(* CODESYS project CanOpen.project (continued)
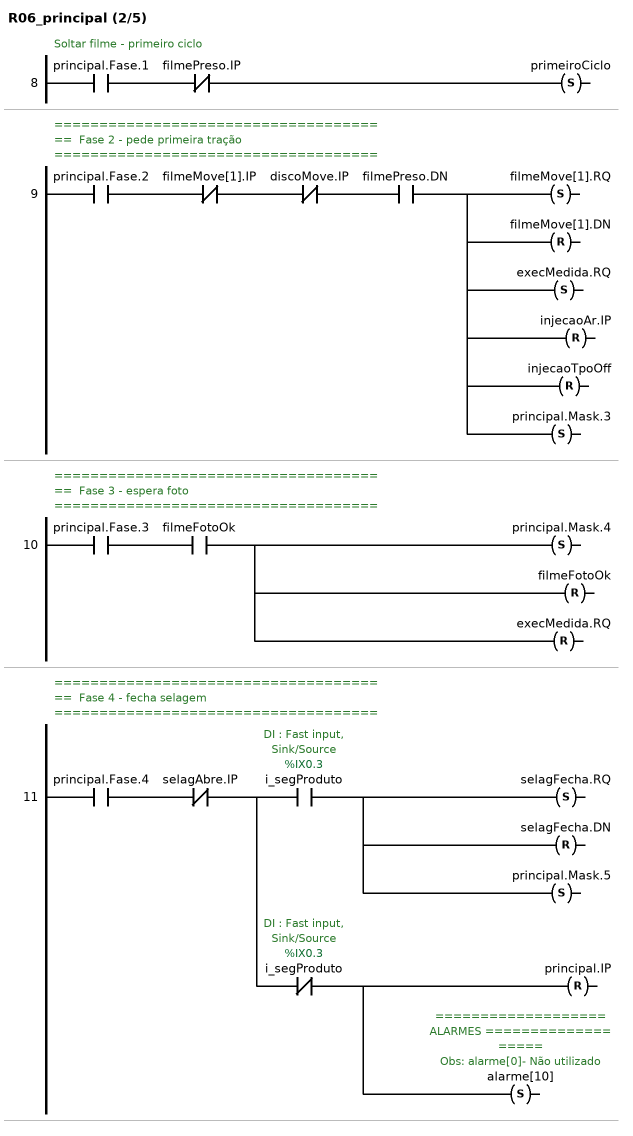
// NETWORK 8
// Soltar filme - primeiro ciclo
primeiroCiclo S= principal.Fase.1 AND NOT filmePreso.IP;

// NETWORK 9
// ====================================
// ==  Fase 2 - pede primeira tração
// ====================================
_w6 := principal.Fase.2 AND NOT filmeMove[1].IP AND NOT discoMove.IP AND filmePreso.DN;
filmeMove[1].RQ S= _w6;
filmeMove[1].DN R= _w6;
execMedida.RQ S= _w6;
injecaoAr.IP R= _w6;
injecaoTpoOff R= _w6;
principal.Mask.3 S= _w6;

// NETWORK 10
// ====================================
// ==  Fase 3 - espera foto
// ====================================
_w7 := principal.Fase.3 AND filmeFotoOk;
principal.Mask.4 S= _w7;
filmeFotoOk R= _w7;
execMedida.RQ R= _w7;

// NETWORK 11
// ====================================
// ==  Fase 4 - fecha selagem
// ====================================
//   i_segProduto: DI : Fast input, Sink/Source | AT %IX0.3
//   alarme[10]: =================== ALARMES =================== Obs: alarme[0]- Não utilizado
_w8 := principal.Fase.4 AND NOT selagAbre.IP;
_w9 := _w8 AND i_segProduto;
selagFecha.RQ S= _w9;
selagFecha.DN R= _w9;
principal.Mask.5 S= _w9;
_w10 := _w8 AND NOT i_segProduto;
principal.IP R= _w10;
alarme[10] S= _w10;

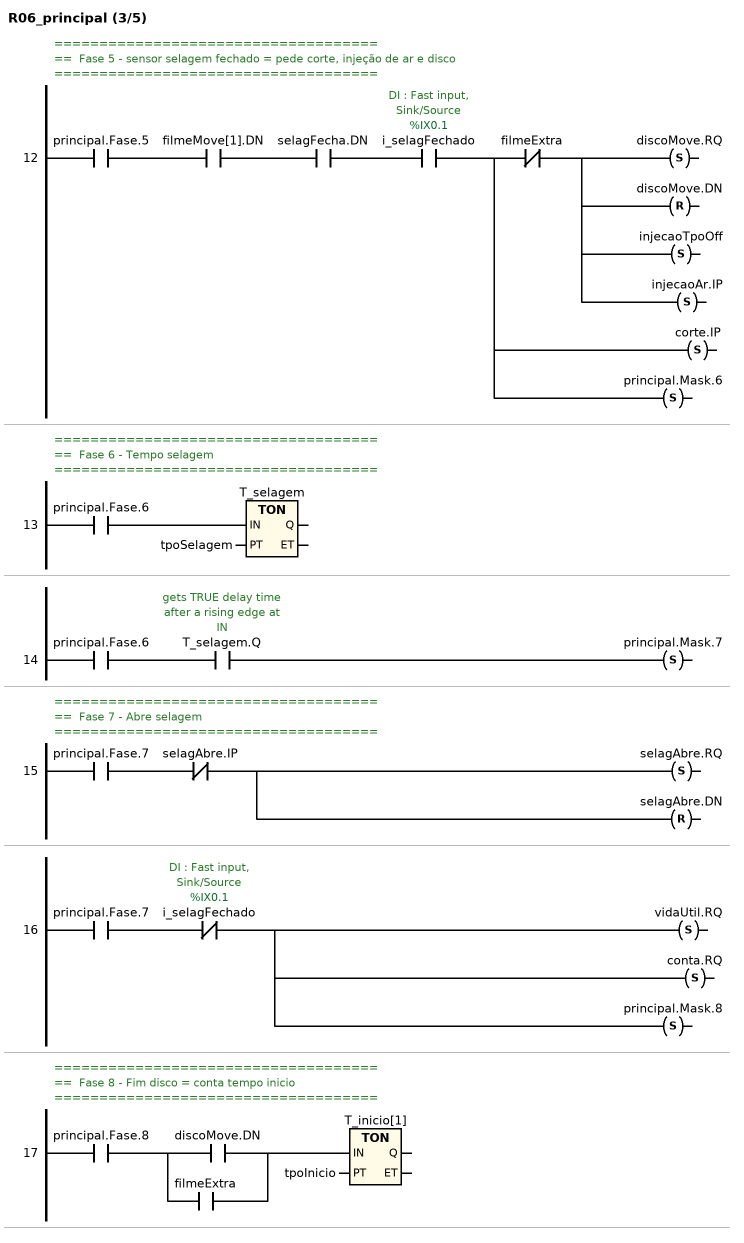
// NETWORK 12
// ====================================
// ==  Fase 5 - sensor selagem fechado = pede corte, injeção de ar e disco
// ====================================
//   i_selagFechado: DI : Fast input, Sink/Source | AT %IX0.1
_w11 := principal.Fase.5 AND filmeMove[1].DN AND selagFecha.DN AND i_selagFechado;
_w12 := _w11 AND NOT filmeExtra;
discoMove.RQ S= _w12;
discoMove.DN R= _w12;
injecaoTpoOff S= _w12;
injecaoAr.IP S= _w12;
corte.IP S= _w11;
principal.Mask.6 S= _w11;

// NETWORK 13
// ====================================
// ==  Fase 6 - Tempo selagem
// ====================================
T_selagem(IN := principal.Fase.6, PT := tpoSelagem); // TON

// NETWORK 14
//   T_selagem.Q: gets TRUE delay time after a rising edge at IN
principal.Mask.7 S= principal.Fase.6 AND T_selagem.Q;

// NETWORK 15
// ====================================
// ==  Fase 7 - Abre selagem
// ====================================
_w13 := principal.Fase.7 AND NOT selagAbre.IP;
selagAbre.RQ S= _w13;
selagAbre.DN R= _w13;

// NETWORK 16
//   i_selagFechado: DI : Fast input, Sink/Source | AT %IX0.1
_w14 := principal.Fase.7 AND NOT i_selagFechado;
vidaUtil.RQ S= _w14;
conta.RQ S= _w14;
principal.Mask.8 S= _w14;

// NETWORK 17
// ====================================
// ==  Fase 8 - Fim disco = conta tempo inicio
// ====================================
T_inicio[1](IN := principal.Fase.8 AND (discoMove.DN OR filmeExtra), PT := tpoInicio); // TON

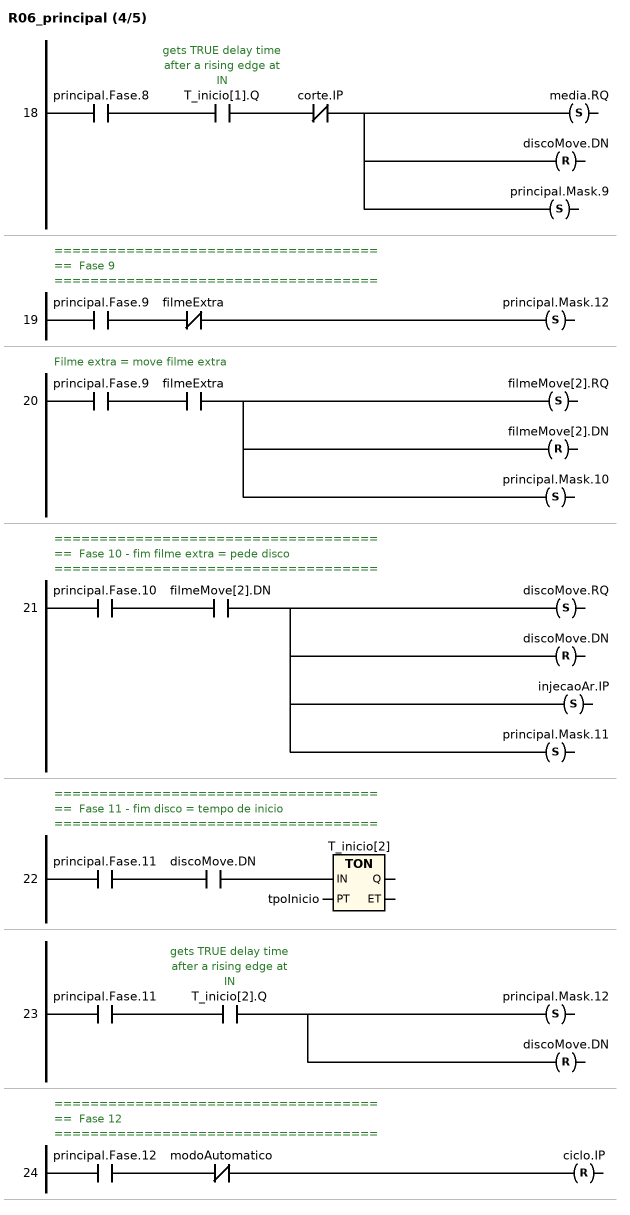
// NETWORK 18
//   T_inicio[1].Q: gets TRUE delay time after a rising edge at IN
_w15 := principal.Fase.8 AND T_inicio[1].Q AND NOT corte.IP;
media.RQ S= _w15;
discoMove.DN R= _w15;
principal.Mask.9 S= _w15;

// NETWORK 19
// ====================================
// ==  Fase 9
// ====================================
principal.Mask.12 S= principal.Fase.9 AND NOT filmeExtra;

// NETWORK 20
// Filme extra = move filme extra
_w16 := principal.Fase.9 AND filmeExtra;
filmeMove[2].RQ S= _w16;
filmeMove[2].DN R= _w16;
principal.Mask.10 S= _w16;

// NETWORK 21
// ====================================
// ==  Fase 10 - fim filme extra = pede disco
// ====================================
_w17 := principal.Fase.10 AND filmeMove[2].DN;
discoMove.RQ S= _w17;
discoMove.DN R= _w17;
injecaoAr.IP S= _w17;
principal.Mask.11 S= _w17;

// NETWORK 22
// ====================================
// ==  Fase 11 - fim disco = tempo de inicio
// ====================================
T_inicio[2](IN := principal.Fase.11 AND discoMove.DN, PT := tpoInicio); // TON

// NETWORK 23
//   T_inicio[2].Q: gets TRUE delay time after a rising edge at IN
_w18 := principal.Fase.11 AND T_inicio[2].Q;
principal.Mask.12 S= _w18;
discoMove.DN R= _w18;

// NETWORK 24
// ====================================
// ==  Fase 12
// ====================================
ciclo.IP R= principal.Fase.12 AND NOT modoAutomatico;

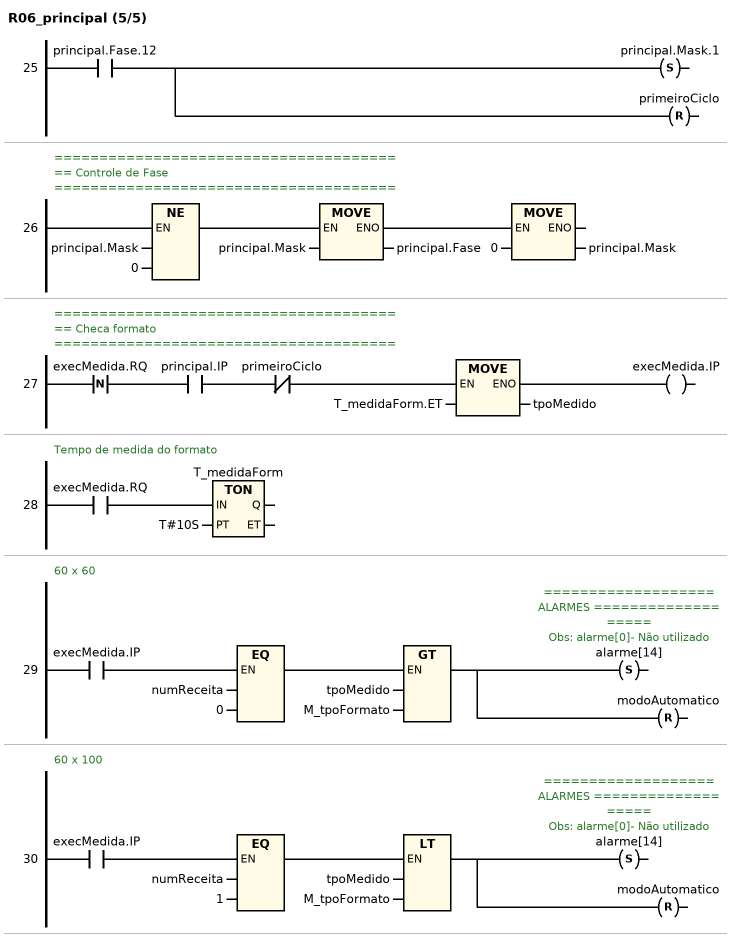
// NETWORK 25
_w19 := principal.Fase.12;
principal.Mask.1 S= _w19;
primeiroCiclo R= _w19;

// NETWORK 26
// ======================================
// == Controle de Fase
// ======================================
_w20 := principal.Mask <> 0;
IF _w20 THEN principal.Fase := principal.Mask; END_IF
IF _w20 THEN principal.Mask := 0; END_IF

// NETWORK 27
// ======================================
// == Checa formato
// ======================================
//   T_medidaForm.ET: elapsed time since rising edge at IN
_ft2(CLK := execMedida.RQ);
_w21 := _ft2.Q AND principal.IP AND NOT primeiroCiclo;
IF _w21 THEN tpoMedido := T_medidaForm.ET; END_IF
execMedida.IP := _w21;

// NETWORK 28
// Tempo de medida do formato
T_medidaForm(IN := execMedida.RQ, PT := T#10S); // TON

// NETWORK 29
// 60 x 60
//   alarme[14]: =================== ALARMES =================== Obs: alarme[0]- Não utilizado
_w22 := execMedida.IP AND numReceita = 0 AND tpoMedido > M_tpoFormato;
alarme[14] S= _w22;
modoAutomatico R= _w22;

// NETWORK 30
// 60 x 100
//   alarme[14]: =================== ALARMES =================== Obs: alarme[0]- Não utilizado
_w23 := execMedida.IP AND numReceita = 1 AND tpoMedido < M_tpoFormato;
alarme[14] S= _w23;
modoAutomatico R= _w23;

END_PROGRAM

// MyController/Application/01_Machine/R21_estatistica
PROGRAM R21_estatistica
VAR
	infoTpoEnergizado			: RTO;
	infoTpoProducao				: RTO;
	auxHrsMinEnerg				: REAL;
	auxHrsMinProd				: REAL;				
END_VAR

(*====================================
  ==  Tempo energizado
  ====================================*)
infoTpoEnergizado(IN:= TRUE,
	  			  PT:= T#60S);
				  
infoTpoEnergizado.RST:= FALSE;			  
IF infoTpoEnergizado.Q THEN
	infoTpoEnergMin:= infoTpoEnergMin + 1;
	IF infoTpoEnergMin > 59 THEN
		infoTpoEnergHrs:= infoTpoEnergHrs + 1;
		infoTpoEnergMin:= 0;
	END_IF
	
	infoTpoEnergizado.RST:= TRUE;
END_IF


(*====================================
  ==  Tempo em produção
  ====================================*)
infoTpoProducao(IN:= ciclo.IP,
	  			PT:= T#60S);
				
IF infoTpoProducao.Q THEN
	infoTpoProdMin:= infoTpoProdMin + 1;
	IF infoTpoProdMin > 59 THEN
		infoTpoProdHrs:= infoTpoProdHrs + 1;
		infoTpoProdMin:= 0;
	END_IF
	
	infoTpoProducao.RST:= TRUE;
END_IF


// Reset dos tempos
IF estatReset THEN
	infoTpoEnergHrs:= 0;
	infoTpoEnergMin:= 0;
	infoTpoProdHrs:= 0;
	infoTpoProdMin:= 0;
	infoTpoEnergizado.RST:= TRUE;
	infoTpoProducao.RST:= TRUE;
	estatReset:= FALSE;
END_IF


(*====================================
  ==  Produtividade
  ====================================*)
// Horas e minutos energizados
auxHrsMinEnerg:= 100.0 * infoTpoEnergHrs + ((100.0 * infoTpoEnergMin) / 60.0);

// Horas e minutos em produção
auxHrsMinProd:= 100.0 * infoTpoProdHrs + ((100.0 * infoTpoProdMin) / 60.0);

IF auxHrsMinEnerg = 0 THEN
	ihm_produtMedio:= 0;
ELSE
	ihm_produtMedio:= (100.0 * auxHrsMinProd) / auxHrsMinEnerg;
END_IF



(*====================================
  ==  Conta
  ====================================*)
// Conta atual e geral
IF conta.RQ THEN
	contaAtual:= contaAtual + 1;
	contaGeral:= contaGeral + 1;
	conta.RQ:= FALSE;
END_IF

// Conta atual maior que programada = gera alarme e parada
IF contaSet <> 0 THEN
	IF contaAtual >= contaSet THEN
		alarme[3]:= TRUE;
		modoAutomatico:= FALSE;
	END_IF
END_IF


// Reset contagem atual
IF contaReset THEN
	contaAtual:= 0;
	contaReset:= FALSE;
END_IF

ihm_contaAtual:= contaAtual;
ihm_contaGeral:= contaGeral;

END_PROGRAM

// MyController/Application/11_FB/RTO
FUNCTION_BLOCK RTO
VAR_INPUT
	IN				: BOOL;
	PT				: TIME;
	RST				: BOOL;
END_VAR
VAR_OUTPUT
	Q				: BOOL;
	ACC				: TIME;
END_VAR
VAR
	auxIn			: BOOL;
	auxAcc			: TIME;
	timer			: TON;
END_VAR

IF IN AND NOT Q THEN
    ACC:= auxAcc + timer.ET;
    auxIn:= true;
end_if;

if not IN then
    auxAcc:= ACC;
    auxIn:= false;
end_if;

if ACC >= PT then
    Q:= true;
    ACC:= PT;
    auxIn:= false;
end_if;

if RST then
    Q:= false;
    ACC:= T#0s;
    auxAcc:= T#0s;
    auxIn:= false;
end_if;

timer(IN:= auxIn, PT:= T#999999S);

END_FUNCTION_BLOCK

// MyController/Application/01_Machine/R22_velocMedia
PROGRAM R22_velocMedia
VAR
	auxVelocMedia			: DINT;
	ctCiclos				: SINT;
	mediaTab				: ARRAY[0..5] OF DINT;
	mediaTpoCiclo			: DINT;
	p0						: SINT;
	T_media					: TON;
	xtr						: ARRAY[0..2] OF R_TRIG;
END_VAR

xtr[0](CLK:= compressor.DN);

IF xtr[0].Q THEN
	ctCiclos:= 0;
END_IF

media.IP:= FALSE;
IF media.RQ THEN
	mediaTpoCiclo:= TIME_TO_DINT(T_media.ET);
	media.RQ:= FALSE;
	media.IP:= TRUE;
END_IF

T_media(IN := compressor.DN AND NOT media.IP,
		PT:= T#600S);

// Carrega valores dentro da tabela		
IF media.IP THEN
	FOR p0:= 1 TO 5 DO
		mediaTab[p0 - 1]:= mediaTab[p0];
	END_FOR
	mediaTab[5]:= mediaTpoCiclo;
	
	// contagem de ciclos para efetuar a média
	IF ctCiclos < 5 THEN
		ctCiclos:= ctCiclos + 1;
	END_IF
	
	
	// Calcula média da tabela
	IF ctCiclos >= 5 THEN
		FOR p0:= 1 TO 5 DO
			IF p0 = 1 THEN
				auxVelocMedia:= 0;  // zera valor no inicio
			END_IF
			 
			auxVelocMedia:= auxVelocMedia + mediaTab[p0]; // soma todos os valores da tabela
		END_FOR
		auxVelocMedia:= auxVelocMedia / 5;
	END_IF
	
	IF auxVelocMedia <> 0 THEN
		ihm_velocMedida:= 60000 / auxVelocMedia;
	END_IF

END_IF;

END_PROGRAM

// MyController/Application/01_Machine/R98_paramFab
PROGRAM R98_paramFab
VAR
END_VAR

paramFab:= FALSE;

(*====================================
  ==  60 x 60
  ====================================*)
 Fb[0].filmeMmAposFoto:= 24;
 Fb[0].discoMmAposFoto:= 0;
 Fb[0].inicioAtraso:= 25;
 Fb[0].discoAtraso:= 20;
 Fb[0].filmeExtra:= FALSE;
 Fb[0].filmeMmExtra:= 1;
 
 
(*====================================
  ==  60 x 100
  ====================================*)
 Fb[1].filmeMmAposFoto:= 24;
 Fb[1].discoMmAposFoto:= 0;
 Fb[1].inicioAtraso:= 25;
 Fb[1].discoAtraso:= 10;
 Fb[1].filmeExtra:= FALSE;
 Fb[1].filmeMmExtra:= 1;
 
 
(*====================================
  ==  70 x 130
  ====================================*)
 Fb[2].filmeMmAposFoto:= 16;
 Fb[2].discoMmAposFoto:= 0;
 Fb[2].inicioAtraso:= 25;
 Fb[2].discoAtraso:= 0;
 Fb[2].filmeExtra:= TRUE;
 Fb[2].filmeMmExtra:= 35;
 
 
(*====================================
  ==  X x Y
  ====================================*)
 Fb[3].filmeMmAposFoto:= 0;
 Fb[3].discoMmAposFoto:= 0;
 Fb[3].inicioAtraso:= 10;
 Fb[3].discoAtraso:= 0;
 Fb[3].filmeExtra:= TRUE;
 Fb[3].filmeMmExtra:= 1;

END_PROGRAM

// MyController/Application/01_Machine/R99_calcTempos
PROGRAM R99_calcTempos
VAR
END_VAR

calcTempos:= FALSE;

// Limita os parametros de atraso de início para 10
IF Fb[numReceita].inicioAtraso < 10 THEN
	Fb[numReceita].inicioAtraso:= 10;
END_IF

IF Rc[numReceita].inicioAtraso < 10 THEN
	Rc[numReceita].inicioAtraso:= 10;
END_IF 

// Cálculo dos tempos
tpoInicio:= DINT_TO_TIME(Rc[numReceita].inicioAtraso) * 10;

tpoDisco:= DINT_TO_TIME(Rc[numReceita].discoAtraso)* 10;

tpoSelagem:= DINT_TO_TIME(M_selagTpoSelagem)* 10;

tpoInjecao:= DINT_TO_TIME(M_tpoInjecaoAr) * 10;

END_PROGRAM

// MyController/Application/02_Filme/F01_geral
PROGRAM F01_geral
VAR
	TD_power				: TOF;
END_VAR

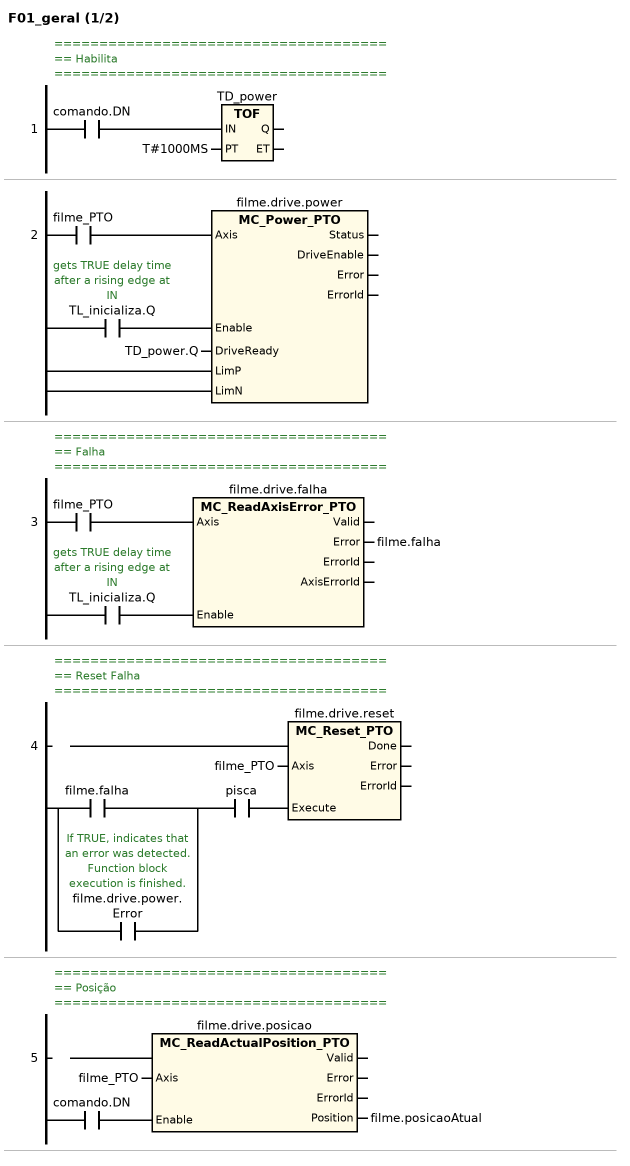
// NETWORK 1
// =====================================
// == Habilita
// =====================================
TD_power(IN := comando.DN, PT := T#1000MS); // TOF

// NETWORK 2
//   TL_inicializa.Q: gets TRUE delay time after a rising edge at IN
//   TD_power.Q: gets FALSE, when PT milliseconds elapsed, since falling edge at IN
filme.drive.power(
    Axis := filme_PTO,
    Enable := TL_inicializa.Q,
    DriveReady := TD_power.Q,
    LimP := TRUE,
    LimN := TRUE); // MC_Power_PTO

// NETWORK 3
// =====================================
// == Falha
// =====================================
//   TL_inicializa.Q: gets TRUE delay time after a rising edge at IN
filme.drive.falha(Axis := filme_PTO, Enable := TL_inicializa.Q, Error => filme.falha); // MC_ReadAxisError_PTO

// NETWORK 4
// =====================================
// == Reset Falha
// =====================================
//   filme.drive.power.Error: If TRUE, indicates that an error was detected. Function block execution is finished.
filme.drive.reset(Axis := filme_PTO, Execute := (filme.falha OR filme.drive.power.Error) AND pisca); // MC_Reset_PTO

// NETWORK 5
// =====================================
// == Posição
// =====================================
filme.drive.posicao(Axis := filme_PTO, Enable := comando.DN, Position => filme.posicaoAtual); // MC_ReadActualPosition_PTO

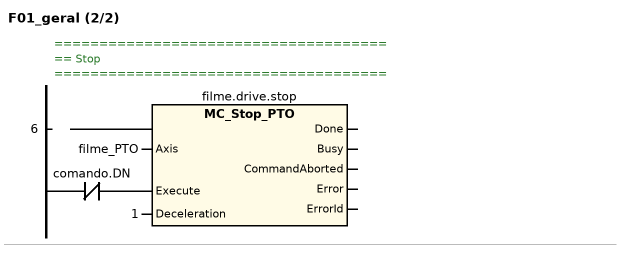
// NETWORK 6
// =====================================
// == Stop
// =====================================
filme.drive.stop(Axis := filme_PTO, Execute := NOT comando.DN, Deceleration := 1); // MC_Stop_PTO

END_PROGRAM

// MyController/Application/02_Filme/F03_auto
PROGRAM F03_auto
VAR
	TF_foto						: TON;
END_VAR
VAR // added by the converter: edge detectors and wires of the graphical bodies
    _w1, _w2, _w3, _w4 : BOOL;
    _ft1 : F_TRIG;
END_VAR

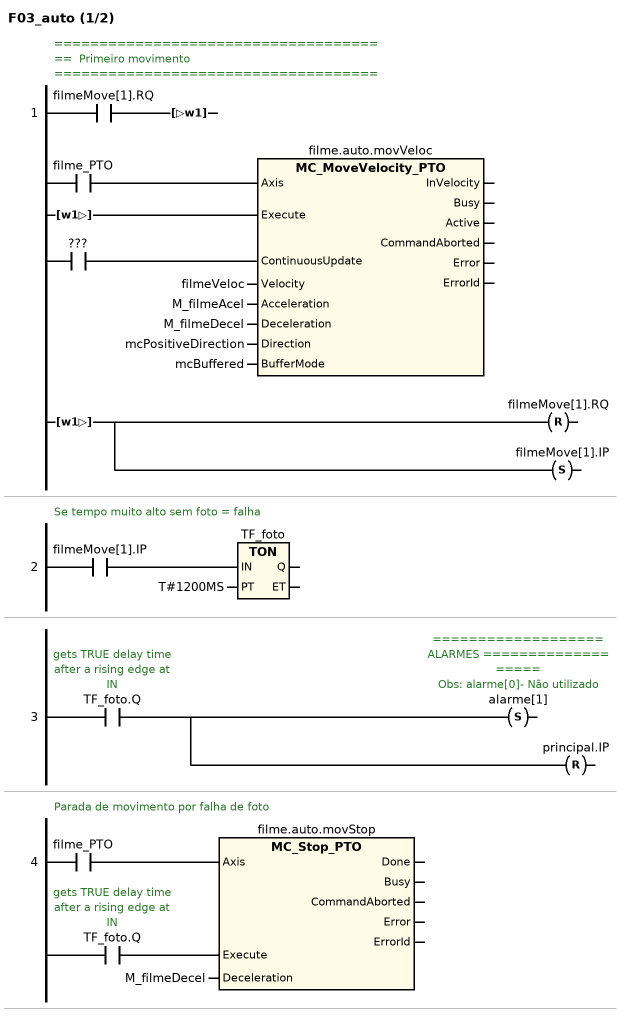
// NETWORK 1
// ====================================
// ==  Primeiro movimento
// ====================================
_w1 := filmeMove[1].RQ;
filme.auto.movVeloc(
    Axis := filme_PTO,
    Execute := _w1,
    Velocity := filmeVeloc,
    Acceleration := M_filmeAcel,
    Deceleration := M_filmeDecel,
    Direction := mcPositiveDirection,
    BufferMode := mcBuffered); // MC_MoveVelocity_PTO
filmeMove[1].RQ R= _w1;
filmeMove[1].IP S= _w1;

// NETWORK 2
// Se tempo muito alto sem foto = falha
TF_foto(IN := filmeMove[1].IP, PT := T#1200MS); // TON

// NETWORK 3
//   TF_foto.Q: gets TRUE delay time after a rising edge at IN
//   alarme[1]: =================== ALARMES =================== Obs: alarme[0]- Não utilizado
alarme[1] S= TF_foto.Q;
principal.IP R= TF_foto.Q;

// NETWORK 4
// Parada de movimento por falha de foto
//   TF_foto.Q: gets TRUE delay time after a rising edge at IN
filme.auto.movStop(Axis := filme_PTO, Execute := TF_foto.Q, Deceleration := M_filmeDecel); // MC_Stop_PTO

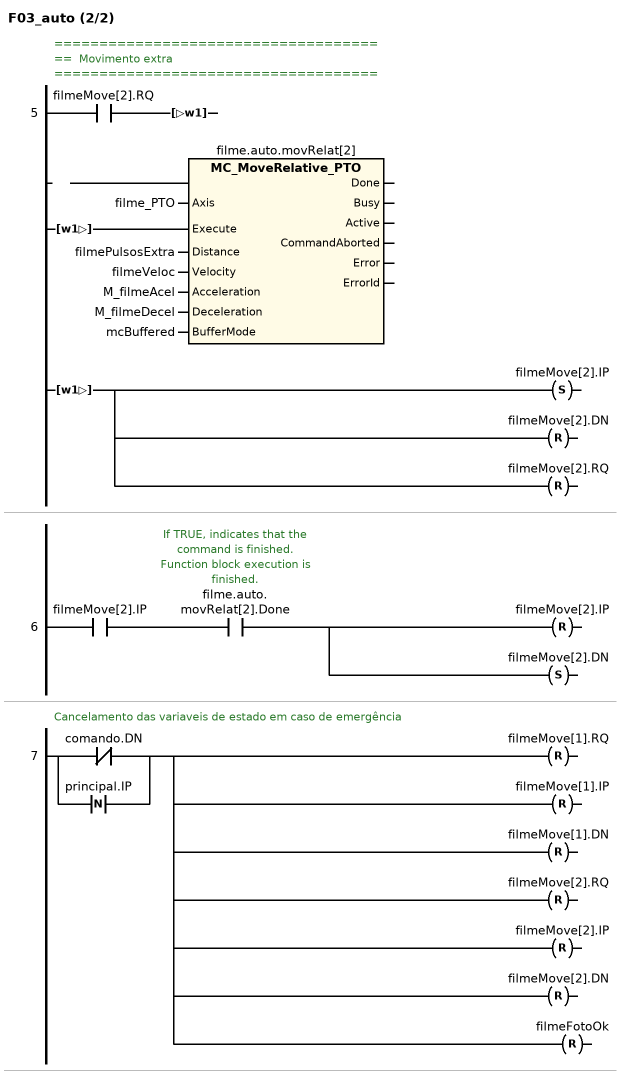
// NETWORK 5
// ====================================
// ==  Movimento extra
// ====================================
_w2 := filmeMove[2].RQ;
filme.auto.movRelat[2](
    Axis := filme_PTO,
    Execute := _w2,
    Distance := filmePulsosExtra,
    Velocity := filmeVeloc,
    Acceleration := M_filmeAcel,
    Deceleration := M_filmeDecel,
    BufferMode := mcBuffered); // MC_MoveRelative_PTO
filmeMove[2].IP S= _w2;
filmeMove[2].DN R= _w2;
filmeMove[2].RQ R= _w2;

// NETWORK 6
//   filme.auto.movRelat[2].Done: If TRUE, indicates that the command is finished. Function block execution is finished.
_w3 := filmeMove[2].IP AND filme.auto.movRelat[2].Done;
filmeMove[2].IP R= _w3;
filmeMove[2].DN S= _w3;

// NETWORK 7
// Cancelamento das variaveis de estado em caso de emergência
_ft1(CLK := principal.IP);
_w4 := NOT comando.DN OR _ft1.Q;
filmeMove[1].RQ R= _w4;
filmeMove[1].IP R= _w4;
filmeMove[1].DN R= _w4;
filmeMove[2].RQ R= _w4;
filmeMove[2].IP R= _w4;
filmeMove[2].DN R= _w4;
filmeFotoOk R= _w4;

END_PROGRAM

// MyController/Application/02_Filme/F99_calculo
PROGRAM F99_calculo
VAR
END_VAR

filme.calcula:= FALSE;

// Limita os parametros de pulsos extra para 1
IF Fb[numReceita].filmeMmExtra < 1 THEN
	Fb[numReceita].filmeMmExtra:= 1;
END_IF

IF Rc[numReceita].filmeMmExtra < 1 THEN
	Rc[numReceita].filmeMmExtra:= 1;
END_IF

// cálculo do num pulsos/mm
filmePulsosMm:= DINT_TO_REAL(M_filmePulsosVolta) / (pi * M_diamRolo);

// cálculo das distâncias a serem percorridas
filmePulsosAposFoto:= REAL_TO_DINT(Rc[numReceita].filmeMmAposFoto * filmePulsosMm);

IF filmePulsosAposFoto = 0 THEN
	filmePulsosAposFoto:= 4;
END_IF

filmePulsosExtra:= REAL_TO_DINT(Rc[numReceita].filmeMmExtra * filmePulsosMm);

// cálculo da velocidade
filmeVeloc:= 350 * M_filmePulsosVolta * M_filmeVeloc / 6000;

END_PROGRAM

// MyController/Application/03_Selagem/S01_geral
PROGRAM S01_geral
VAR
	TD_power			: TOF;
END_VAR
VAR // added by the converter: edge detectors and wires of the graphical bodies
    _ft1 : F_TRIG;
END_VAR

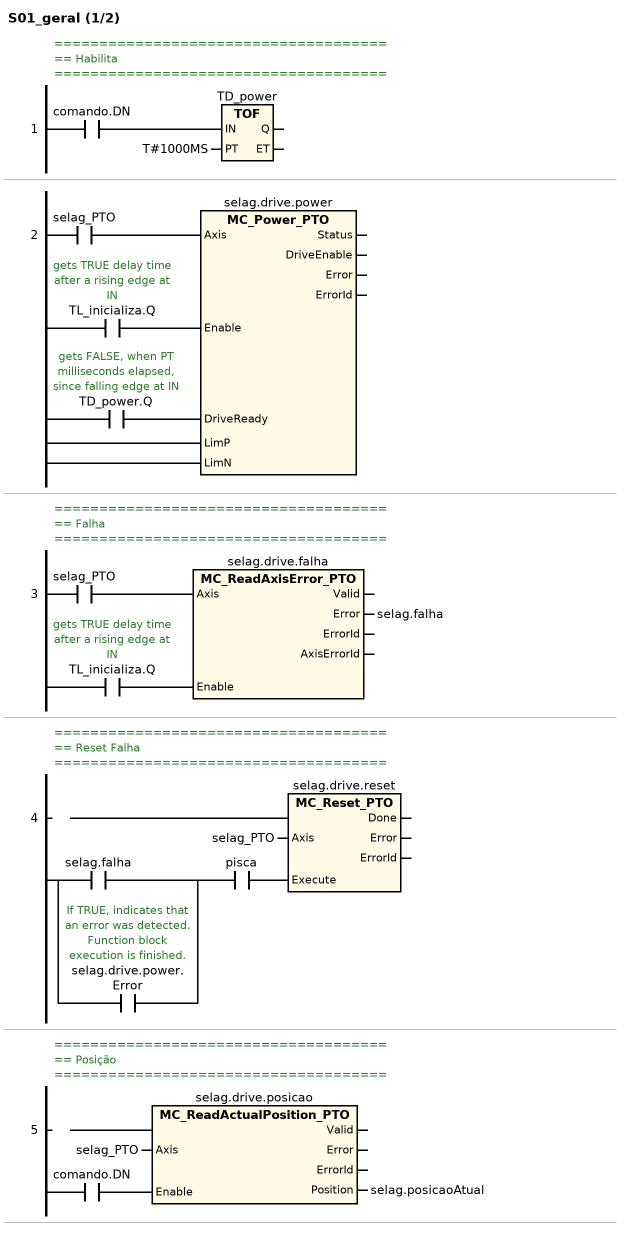
// NETWORK 1
// =====================================
// == Habilita
// =====================================
TD_power(IN := comando.DN, PT := T#1000MS); // TOF

// NETWORK 2
//   TL_inicializa.Q: gets TRUE delay time after a rising edge at IN
//   TD_power.Q: gets FALSE, when PT milliseconds elapsed, since falling edge at IN
selag.drive.power(
    Axis := selag_PTO,
    Enable := TL_inicializa.Q,
    DriveReady := TD_power.Q,
    LimP := TRUE,
    LimN := TRUE); // MC_Power_PTO

// NETWORK 3
// =====================================
// == Falha
// =====================================
//   TL_inicializa.Q: gets TRUE delay time after a rising edge at IN
selag.drive.falha(Axis := selag_PTO, Enable := TL_inicializa.Q, Error => selag.falha); // MC_ReadAxisError_PTO

// NETWORK 4
// =====================================
// == Reset Falha
// =====================================
//   selag.drive.power.Error: If TRUE, indicates that an error was detected. Function block execution is finished.
selag.drive.reset(Axis := selag_PTO, Execute := (selag.falha OR selag.drive.power.Error) AND pisca); // MC_Reset_PTO

// NETWORK 5
// =====================================
// == Posição
// =====================================
selag.drive.posicao(Axis := selag_PTO, Enable := comando.DN, Position => selag.posicaoAtual); // MC_ReadActualPosition_PTO

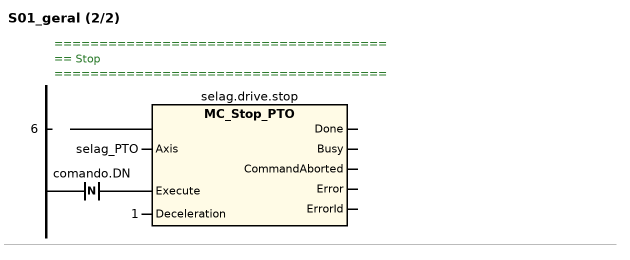
// NETWORK 6
// =====================================
// == Stop
// =====================================
_ft1(CLK := comando.DN);
selag.drive.stop(Axis := selag_PTO, Execute := _ft1.Q, Deceleration := 1); // MC_Stop_PTO

END_PROGRAM

// MyController/Application/03_Selagem/S02_home
PROGRAM S02_home
VAR
	auxDword				: DWORD;
	TF_home					: TON;
END_VAR
VAR // added by the converter: edge detectors and wires of the graphical bodies
    _rt1 : R_TRIG;
    _w1, _w2, _w3, _w4, _w5 : BOOL;
END_VAR

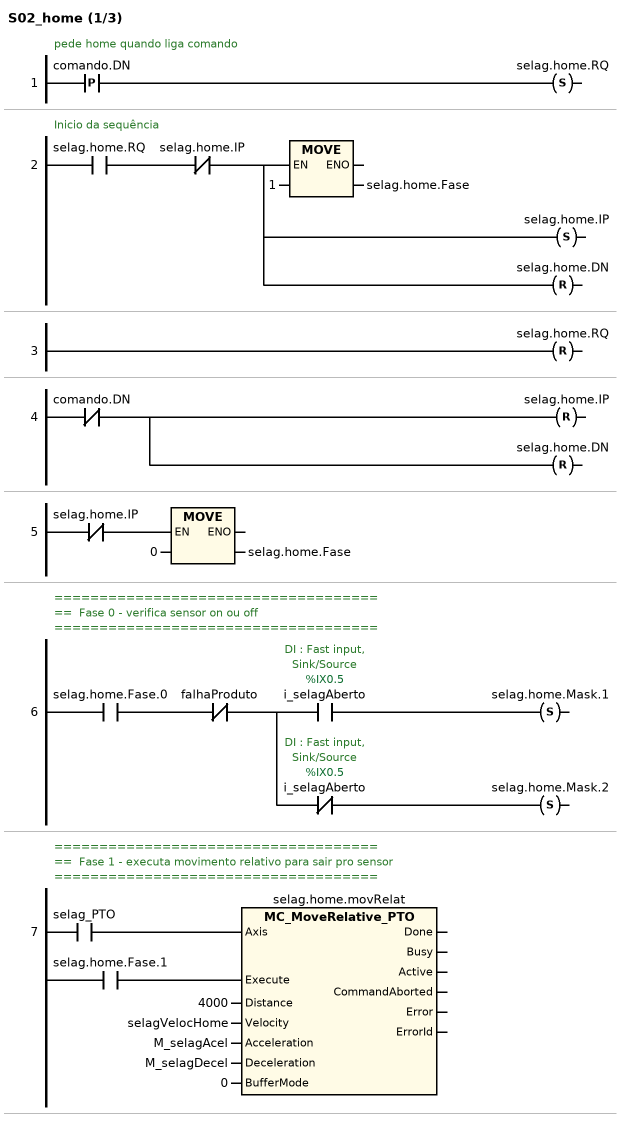
// NETWORK 1
// pede home quando liga comando
_rt1(CLK := comando.DN);
selag.home.RQ S= _rt1.Q;

// NETWORK 2
// Inicio da sequência
_w1 := selag.home.RQ AND NOT selag.home.IP;
IF _w1 THEN selag.home.Fase := 1; END_IF
selag.home.IP S= _w1;
selag.home.DN R= _w1;

// NETWORK 3
selag.home.RQ R= TRUE;

// NETWORK 4
_w2 := NOT comando.DN;
selag.home.IP R= _w2;
selag.home.DN R= _w2;

// NETWORK 5
IF NOT selag.home.IP THEN selag.home.Fase := 0; END_IF

// NETWORK 6
// ====================================
// ==  Fase 0 - verifica sensor on ou off
// ====================================
//   i_selagAberto: DI : Fast input, Sink/Source | AT %IX0.5
_w3 := selag.home.Fase.0 AND NOT falhaProduto;
selag.home.Mask.1 S= _w3 AND i_selagAberto;
selag.home.Mask.2 S= _w3 AND NOT i_selagAberto;

// NETWORK 7
// ====================================
// ==  Fase 1 - executa movimento relativo para sair pro sensor
// ====================================
selag.home.movRelat(
    Axis := selag_PTO,
    Execute := selag.home.Fase.1,
    Distance := 4000,
    Velocity := selagVelocHome,
    Acceleration := M_selagAcel,
    Deceleration := M_selagDecel,
    BufferMode := 0); // MC_MoveRelative_PTO

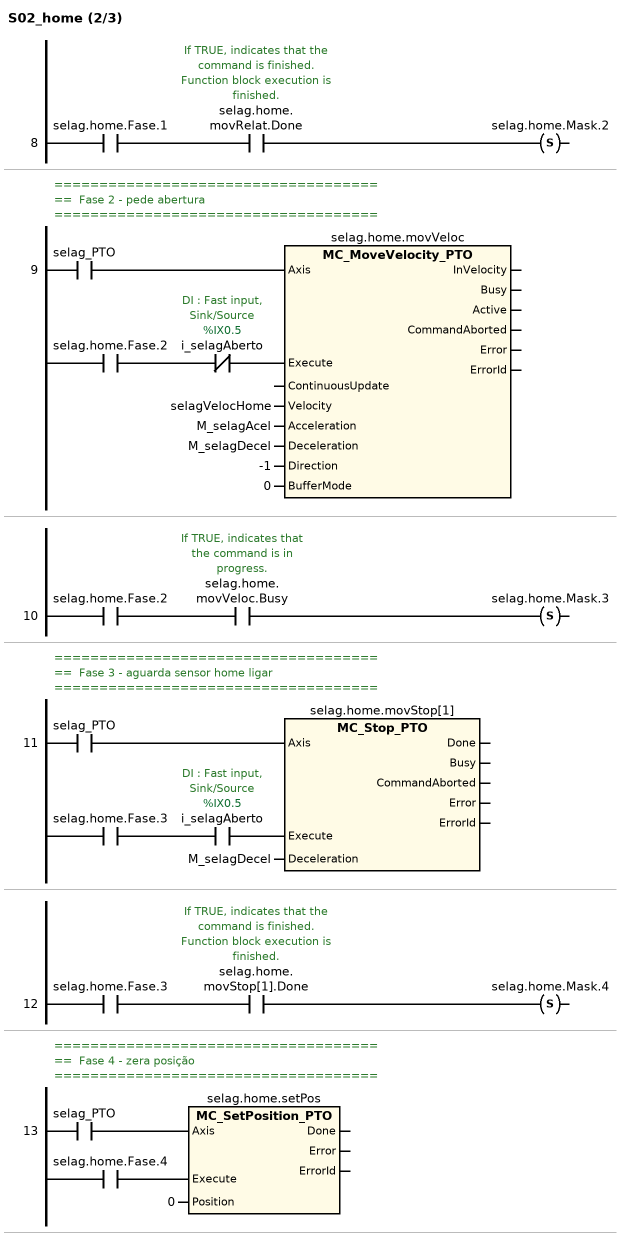
// NETWORK 8
//   selag.home.movRelat.Done: If TRUE, indicates that the command is finished. Function block execution is finished.
selag.home.Mask.2 S= selag.home.Fase.1 AND selag.home.movRelat.Done;

// NETWORK 9
// ====================================
// ==  Fase 2 - pede abertura
// ====================================
//   i_selagAberto: DI : Fast input, Sink/Source | AT %IX0.5
selag.home.movVeloc(
    Axis := selag_PTO,
    Execute := selag.home.Fase.2 AND NOT i_selagAberto,
    Velocity := selagVelocHome,
    Acceleration := M_selagAcel,
    Deceleration := M_selagDecel,
    Direction := -1,
    BufferMode := 0); // MC_MoveVelocity_PTO

// NETWORK 10
//   selag.home.movVeloc.Busy: If TRUE, indicates that the command is in progress.
selag.home.Mask.3 S= selag.home.Fase.2 AND selag.home.movVeloc.Busy;

// NETWORK 11
// ====================================
// ==  Fase 3 - aguarda sensor home ligar
// ====================================
//   i_selagAberto: DI : Fast input, Sink/Source | AT %IX0.5
selag.home.movStop[1](
    Axis := selag_PTO,
    Execute := selag.home.Fase.3 AND i_selagAberto,
    Deceleration := M_selagDecel); // MC_Stop_PTO

// NETWORK 12
//   selag.home.movStop[1].Done: If TRUE, indicates that the command is finished. Function block execution is finished.
selag.home.Mask.4 S= selag.home.Fase.3 AND selag.home.movStop[1].Done;

// NETWORK 13
// ====================================
// ==  Fase 4 - zera posição
// ====================================
selag.home.setPos(Axis := selag_PTO, Execute := selag.home.Fase.4, Position := 0); // MC_SetPosition_PTO

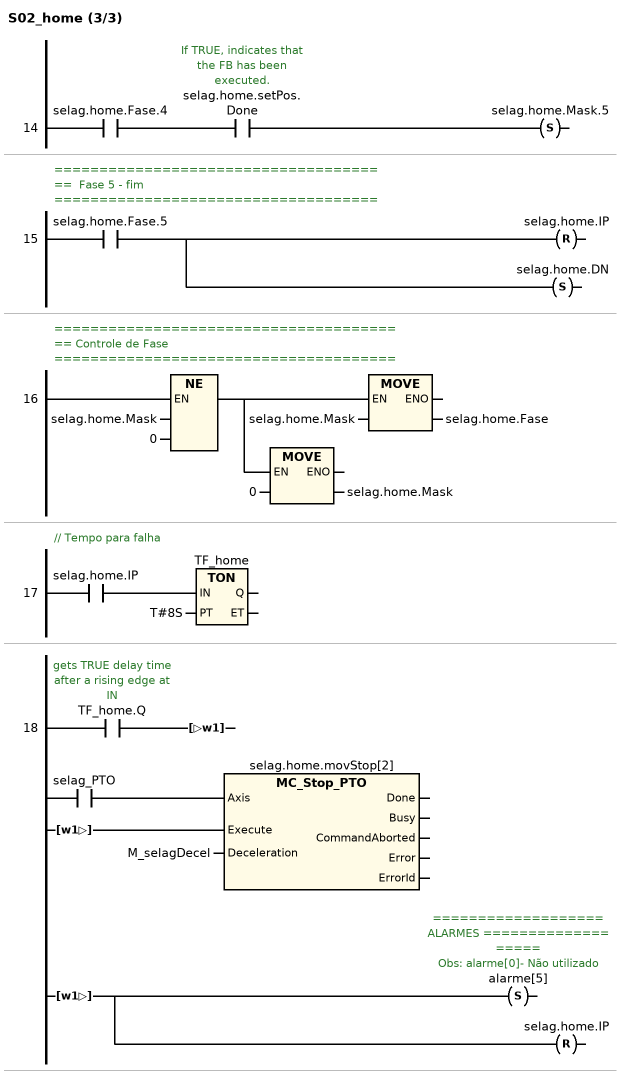
// NETWORK 14
//   selag.home.setPos.Done: If TRUE, indicates that the FB has been executed.
selag.home.Mask.5 S= selag.home.Fase.4 AND selag.home.setPos.Done;

// NETWORK 15
// ====================================
// ==  Fase 5 - fim
// ====================================
_w4 := selag.home.Fase.5;
selag.home.IP R= _w4;
selag.home.DN S= _w4;

// NETWORK 16
// ======================================
// == Controle de Fase
// ======================================
_w5 := selag.home.Mask <> 0;
IF _w5 THEN selag.home.Fase := selag.home.Mask; END_IF
IF _w5 THEN selag.home.Mask := 0; END_IF

// NETWORK 17
// // Tempo para falha
TF_home(IN := selag.home.IP, PT := T#8S); // TON

// NETWORK 18
//   TF_home.Q: gets TRUE delay time after a rising edge at IN
//   alarme[5]: =================== ALARMES =================== Obs: alarme[0]- Não utilizado
selag.home.movStop[2](Axis := selag_PTO, Execute := TF_home.Q, Deceleration := M_selagDecel); // MC_Stop_PTO
alarme[5] S= TF_home.Q;
selag.home.IP R= TF_home.Q;

END_PROGRAM

// MyController/Application/03_Selagem/S03_auto
PROGRAM S03_auto
VAR
	TL_home					: TON;
	TF_selagem				: ARRAY[1..2] OF TON;
END_VAR
VAR // added by the converter: edge detectors and wires of the graphical bodies
    _w1, _w2, _w3, _w4, _w5, _w6, _w7, _w8 : BOOL;
    _ft1 : F_TRIG;
END_VAR

